(* Logix 5000 project; controller FV vendor 1 type 14 code 217 rev 31.11; software revision 31.00; part 12 of 63 *)
(* tags used below, declared in another part *)
   CWD : CHECKWORD_FLAGS;
   FR_B240 : INT[255];   // DEBOUNCE Debounce Flags
   FR_B246 : INT[255];   // V_REVERSE Flags for reversing contol action
   FR_B3 : INT[255];   // BINARY
   FR_FV26_AV07 : PlantItem;   // FV26_AV07
   FR_FV26_ROTO : PlantItem;   // FV26_ROTO
   FR_FV27_AV01 : PlantItem;   // FV27_AV01
   FR_FV27_AV04 : PlantItem;   // FV27_AV04
   FR_FV27_AV05 : PlantItem;   // FV27_AV05
   FR_FV27_AV06 : PlantItem;   // FV27_AV06
   FR_FV27_AV07 : PlantItem;   // FV27_AV07
   FR_FV27_ROTO : PlantItem;   // FV27_ROTO
   FR_FV27_VA01 : PlantItem;   // FV27_VA01
   FR_FV28_AV01 : PlantItem;   // FV28_AV01
   FR_FV28_AV04 : PlantItem;   // FV28_AV04
   FR_FV28_AV05 : PlantItem;   // FV28_AV05
   FR_FV28_AV06 : PlantItem;   // FV28_AV06
   FR_FV28_AV07 : PlantItem;   // FV28_AV07
   FR_FV28_ROTO : PlantItem;   // FV28_ROTO
   FR_FV28_V : PlantItem;   // FV28_V
   FR_FV28_VA01 : PlantItem;   // FV28_VA01
   FR_N10 : INT[265];   // FV_AGING Comms to FV Aging PL C
   FR_N100 : INT[265];   // FV FILLING
   FR_N110 : INT[265];   // GREEN BEER Green Beer Main
   FR_N120 : INT[265];   // YEAST CROP Yeast Cropping Main
   FR_N13 : INT[265];   // MV_ROUTE Comms to MV Routing PLC
   FR_N130 : INT[265];   // FILTRATE Filtrate Return
   FR_N14 : INT[265];   // MVFV CIP Comms to MVFV CIP Un it PLC
   FR_N160 : INT[265];   // VESSEL Vessel Working Direc tory
   FR_N200 : INT[265];   // ANALOG_IN Analog Inputs
   FR_N255 : INT[265];   // CHECKWORDS
   FR_N26 : INT[265];   // FV26
   FR_N27 : INT[265];   // FV27
   FR_N28 : INT[265];   // FV28
   FR_N7 : INT[265];   // INTEGER
   FR_N99 : INT[265];   // COMMENT Comment Lines
   FR_T144 : TIMER[255];   // CIP
   FR_T4 : TIMER[255];   // TIMER
   FR_T50 : TIMER[52];
   FR_T51 : TIMER[52];
   FR_T52 : TIMER[52];
   FR_T53 : TIMER[52];
   FR_VB1_AV08 : PlantItem;   // VB1_AV08
   FR_VB1_AV09 : PlantItem;   // VB1_AV09
   FR_VB2_AV04 : PlantItem;   // VB2_AV04
   FR_VB2_AV05 : PlantItem;   // VB2_AV05
   FR_VB4_AV02 : PlantItem;   // VB4_AV02
   FR_VB4_AV06 : PlantItem;   // VB4_AV06
   FR_VB4_AV08 : PlantItem;   // VB4_AV08
   FR_VB4_AV12 : PlantItem;   // VB4_AV12
   FR_VB4_AV14 : PlantItem;   // VB4_AV14
   FR_VB4_AV18 : PlantItem;   // VB4_AV18
(* FR_Common, continued *)

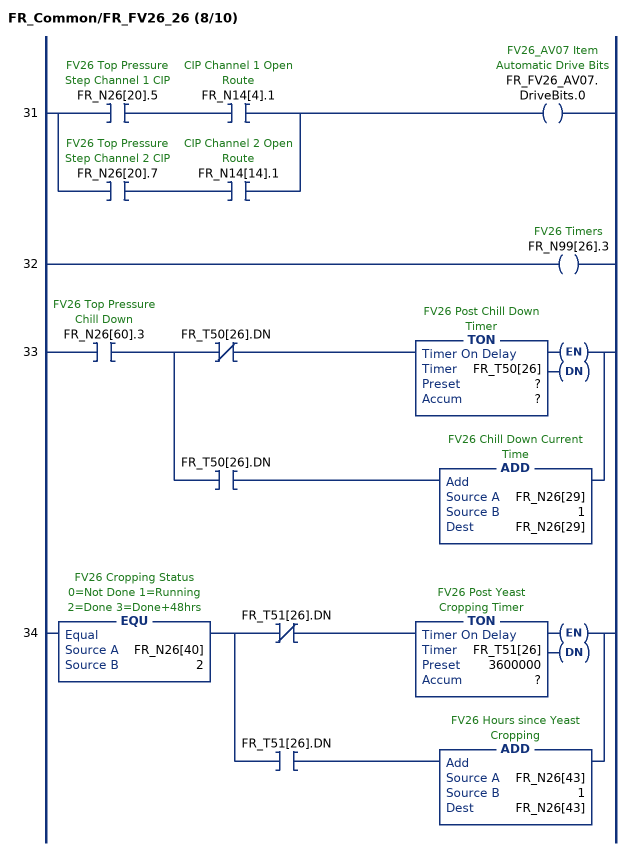
   [picture p160: FR_Common/FR_FV26_26 rungs 31-34]
   31: [XIC(FR_N26[20].5) XIC(FR_N14[4].1) ,XIC(FR_N26[20].7) XIC(FR_N14[14].1) ]OTE(FR_FV26_AV07.DriveBits.0);
   32: OTE(FR_N99[26].3);
   33: XIC(FR_N26[60].3)[XIO(FR_T50[26].DN) TON(FR_T50[26],?,?) ,XIC(FR_T50[26].DN) ADD(FR_N26[29],1,FR_N26[29]) ];
   34: EQU(FR_N26[40],2)[XIO(FR_T51[26].DN) TON(FR_T51[26],?,?) ,XIC(FR_T51[26].DN) ADD(FR_N26[43],1,FR_N26[43]) ];
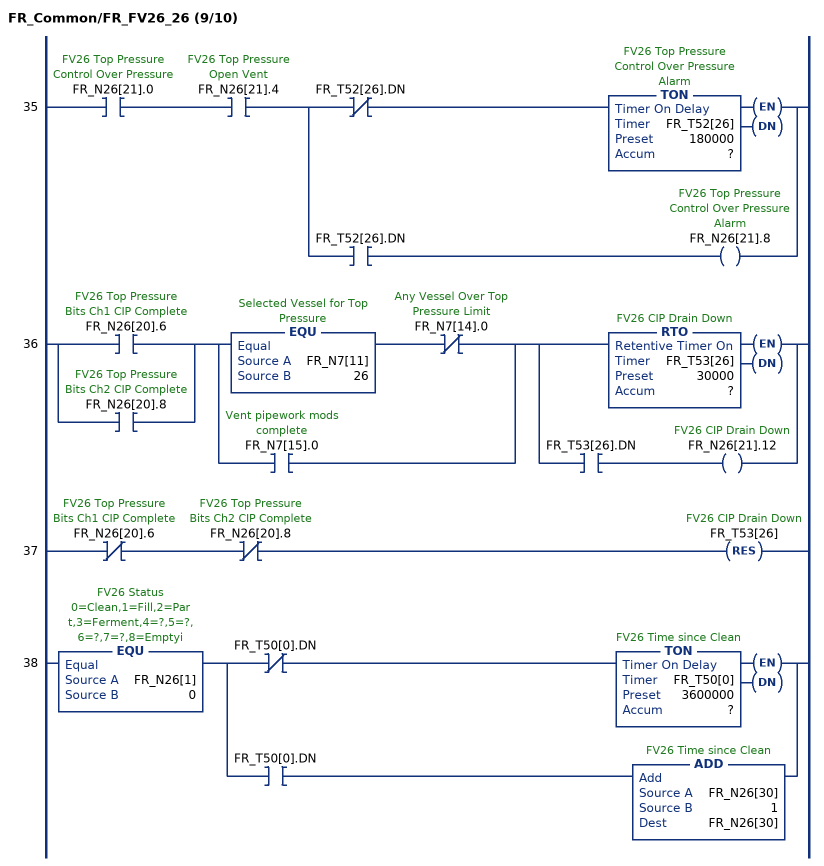
   35: XIC(FR_N26[21].0)XIC(FR_N26[21].4)[XIO(FR_T52[26].DN) TON(FR_T52[26],?,?) ,XIC(FR_T52[26].DN) OTE(FR_N26[21].8) ];
   36: [XIC(FR_N26[20].6) ,XIC(FR_N26[20].8) ][EQU(FR_N7[11],26) XIO(FR_N7[14].0) ,XIC(FR_N7[15].0) ][RTO(FR_T53[26],?,?) ,XIC(FR_T53[26].DN) OTE(FR_N26[21].12) ];
   37: XIO(FR_N26[20].6)XIO(FR_N26[20].8)RES(FR_T53[26]);
   38: EQU(FR_N26[1],0)[XIO(FR_T50[0].DN) TON(FR_T50[0],?,?) ,XIC(FR_T50[0].DN) ADD(FR_N26[30],1,FR_N26[30]) ];
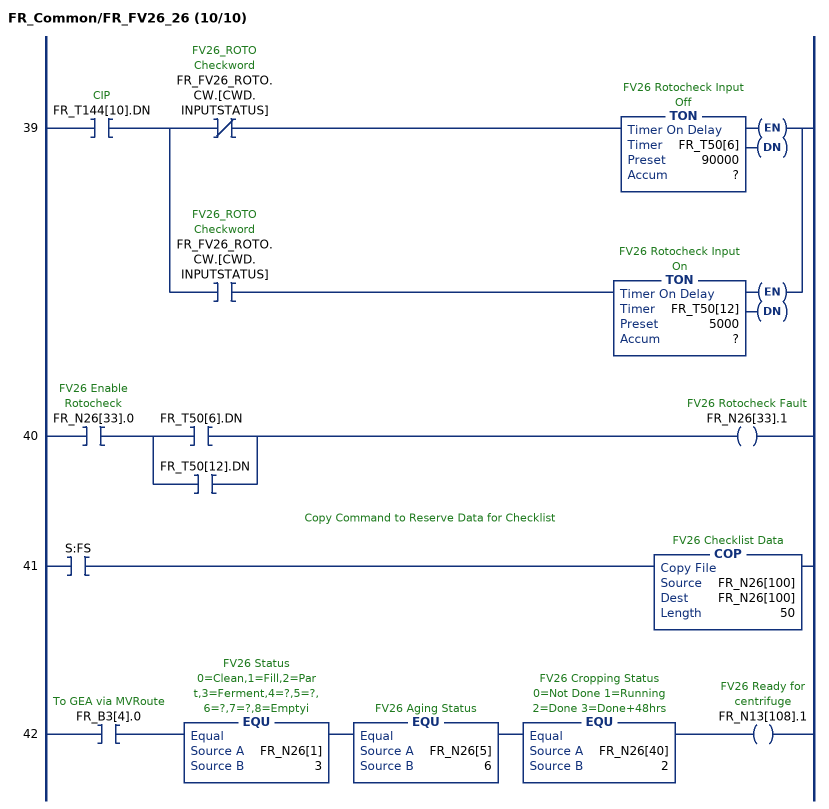
   39: XIC(FR_T144[10].DN)[XIO(FR_FV26_ROTO.CW.[CWD.INPUTSTATUS]) TON(FR_T50[6],?,?) ,XIC(FR_FV26_ROTO.CW.[CWD.INPUTSTATUS]) TON(FR_T50[12],?,?) ];
   40: XIC(FR_N26[33].0)[XIC(FR_T50[6].DN) ,XIC(FR_T50[12].DN) ]OTE(FR_N26[33].1);
   // Copy Command to Reserve Data for Checklist
   41: XIC(S:FS)COP(FR_N26[100],FR_N26[100],50);
   42: XIC(FR_B3[4].0)EQU(FR_N26[1],3)EQU(FR_N26[5],6)EQU(FR_N26[40],2)OTE(FR_N13[108].1);
END_ROUTINE

ROUTINE FR_FV27_27   (* ladder *)
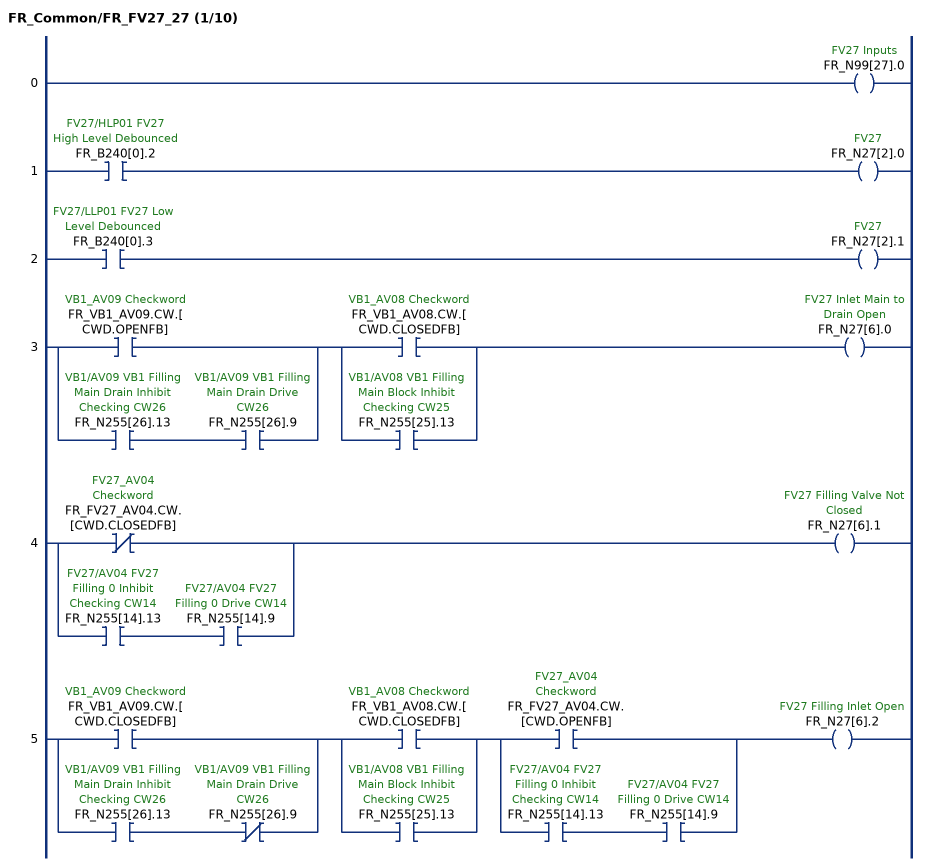
   0: OTE(FR_N99[27].0);
   1: XIC(FR_B240[0].2)OTE(FR_N27[2].0);
   2: XIC(FR_B240[0].3)OTE(FR_N27[2].1);
   3: [XIC(FR_VB1_AV09.CW.[CWD.OPENFB]) ,XIC(FR_N255[26].13) XIC(FR_N255[26].9) ][XIC(FR_VB1_AV08.CW.[CWD.CLOSEDFB]) ,XIC(FR_N255[25].13) ]OTE(FR_N27[6].0);
   4: [XIO(FR_FV27_AV04.CW.[CWD.CLOSEDFB]) ,XIC(FR_N255[14].13) XIC(FR_N255[14].9) ]OTE(FR_N27[6].1);
   5: [XIC(FR_VB1_AV09.CW.[CWD.CLOSEDFB]) ,XIC(FR_N255[26].13) XIO(FR_N255[26].9) ][XIC(FR_VB1_AV08.CW.[CWD.CLOSEDFB]) ,XIC(FR_N255[25].13) ][XIC(FR_FV27_AV04.CW.[CWD.OPENFB]) ,XIC(FR_N255[14].13) XIC(FR_N255[14].9) ]OTE(FR_N27[6].2);
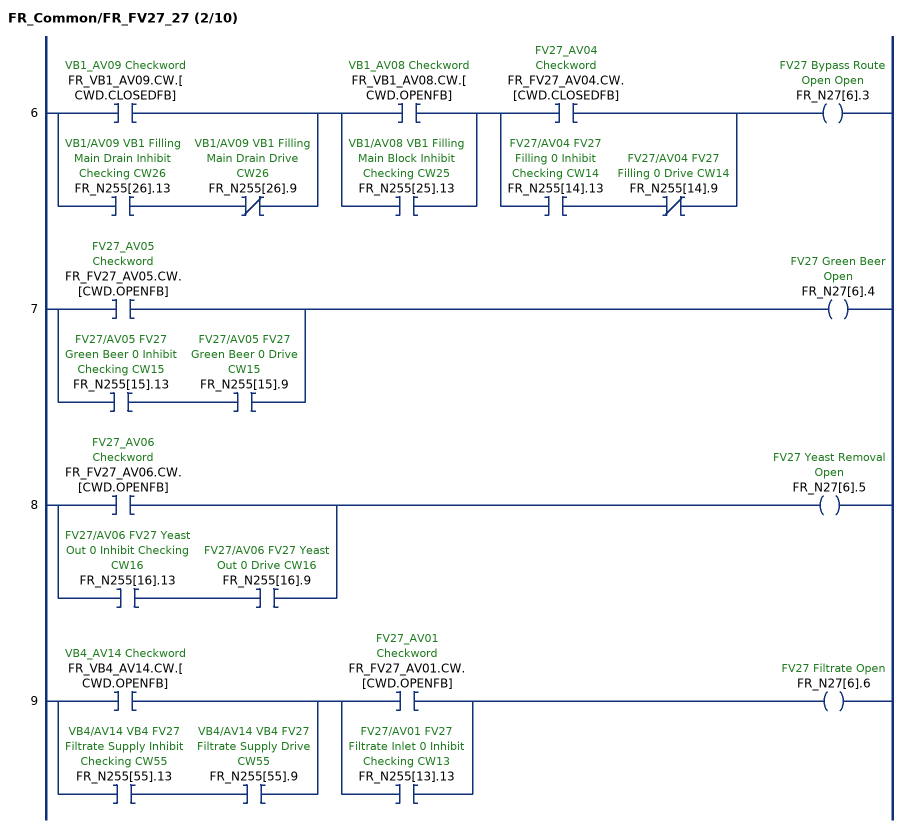
   6: [XIC(FR_VB1_AV09.CW.[CWD.CLOSEDFB]) ,XIC(FR_N255[26].13) XIO(FR_N255[26].9) ][XIC(FR_VB1_AV08.CW.[CWD.OPENFB]) ,XIC(FR_N255[25].13) ][XIC(FR_FV27_AV04.CW.[CWD.CLOSEDFB]) ,XIC(FR_N255[14].13) XIO(FR_N255[14].9) ]OTE(FR_N27[6].3);
   7: [XIC(FR_FV27_AV05.CW.[CWD.OPENFB]) ,XIC(FR_N255[15].13) XIC(FR_N255[15].9) ]OTE(FR_N27[6].4);
   8: [XIC(FR_FV27_AV06.CW.[CWD.OPENFB]) ,XIC(FR_N255[16].13) XIC(FR_N255[16].9) ]OTE(FR_N27[6].5);
   9: [XIC(FR_VB4_AV14.CW.[CWD.OPENFB]) ,XIC(FR_N255[55].13) XIC(FR_N255[55].9) ][XIC(FR_FV27_AV01.CW.[CWD.OPENFB]) ,XIC(FR_N255[13].13) ]OTE(FR_N27[6].6);
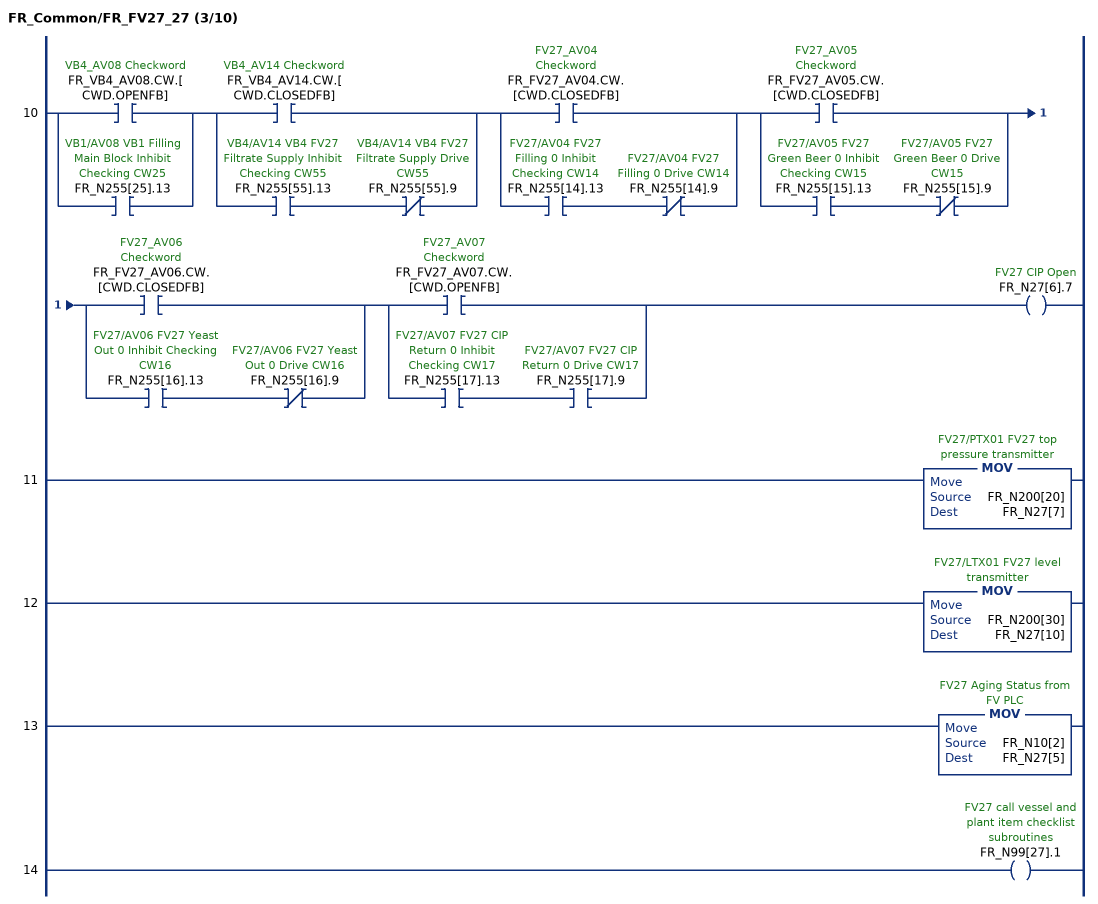
   10: [XIC(FR_VB4_AV08.CW.[CWD.OPENFB]) ,XIC(FR_N255[25].13) ][XIC(FR_VB4_AV14.CW.[CWD.CLOSEDFB]) ,XIC(FR_N255[55].13) XIO(FR_N255[55].9) ][XIC(FR_FV27_AV04.CW.[CWD.CLOSEDFB]) ,XIC(FR_N255[14].13) XIO(FR_N255[14].9) ][XIC(FR_FV27_AV05.CW.[CWD.CLOSEDFB]) ,XIC(FR_N255[15].13) XIO(FR_N255[15].9) ][XIC(FR_FV27_AV06.CW.[CWD.CLOSEDFB]) ,XIC(FR_N255[16].13) XIO(FR_N255[16].9) ][XIC(FR_FV27_AV07.CW.[CWD.OPENFB]) ,XIC(FR_N255[17].13) XIC(FR_N255[17].9) ]OTE(FR_N27[6].7);
   11: MOV(FR_N200[20],FR_N27[7]);
   12: MOV(FR_N200[30],FR_N27[10]);
   13: MOV(FR_N10[2],FR_N27[5]);
   14: OTE(FR_N99[27].1);
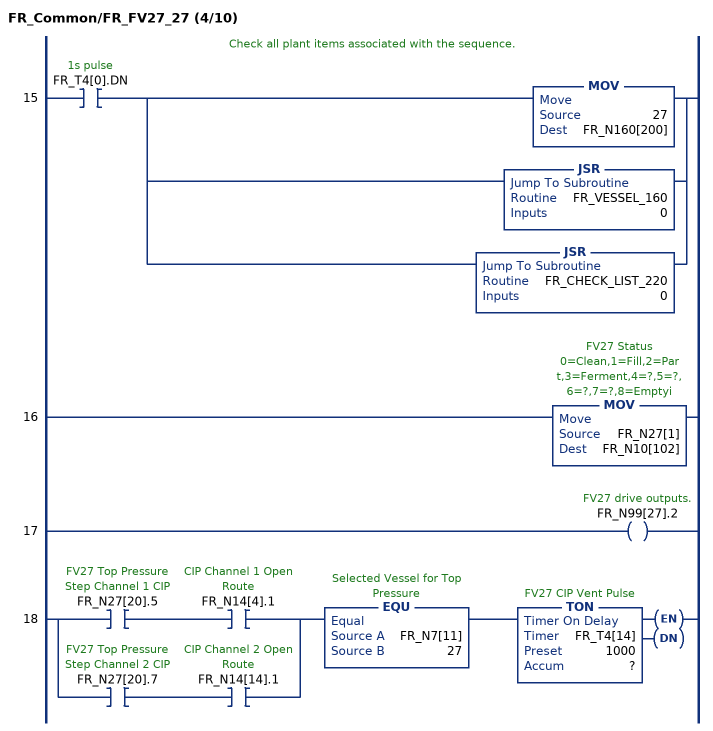
   // Check all plant items associated with the sequence.
   15: XIC(FR_T4[0].DN)[MOV(27,FR_N160[200]) ,JSR(FR_VESSEL_160,0) ,JSR(FR_CHECK_LIST_220,0) ];
   16: MOV(FR_N27[1],FR_N10[102]);
   17: OTE(FR_N99[27].2);
   18: [XIC(FR_N27[20].5) XIC(FR_N14[4].1) ,XIC(FR_N27[20].7) XIC(FR_N14[14].1) ]EQU(FR_N7[11],27)TON(FR_T4[14],?,?);
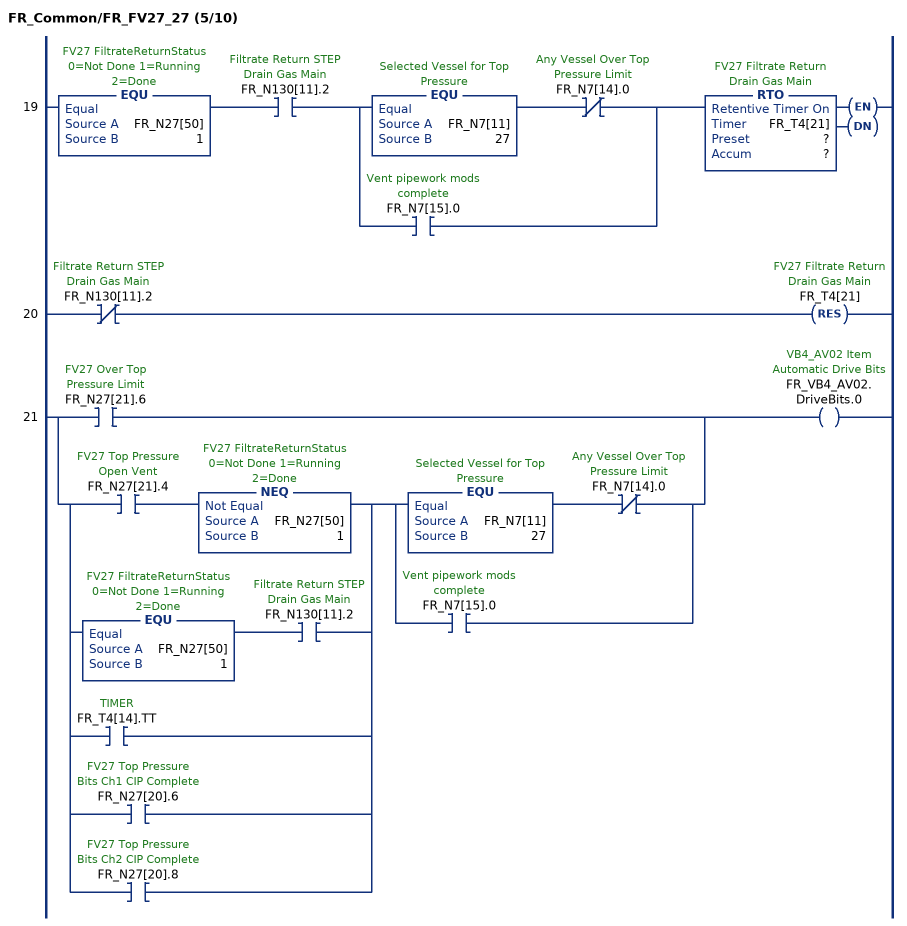
   19: EQU(FR_N27[50],1)XIC(FR_N130[11].2)[EQU(FR_N7[11],27) XIO(FR_N7[14].0) ,XIC(FR_N7[15].0) ]RTO(FR_T4[21],?,?);
   20: XIO(FR_N130[11].2)RES(FR_T4[21]);
   21: [XIC(FR_N27[21].6) ,[XIC(FR_N27[21].4) NEQ(FR_N27[50],1) ,EQU(FR_N27[50],1) XIC(FR_N130[11].2) ,XIC(FR_T4[14].TT) ,[XIC(FR_N27[20].6) ,XIC(FR_N27[20].8) ] ] [EQU(FR_N7[11],27) XIO(FR_N7[14].0) ,XIC(FR_N7[15].0) ] ]OTE(FR_VB4_AV02.DriveBits.0);
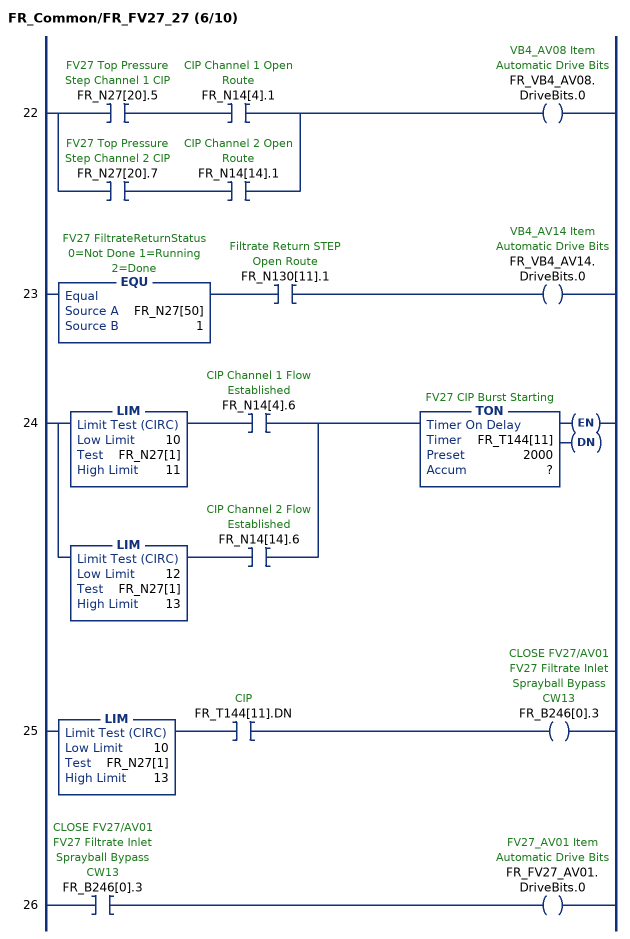
   22: [XIC(FR_N27[20].5) XIC(FR_N14[4].1) ,XIC(FR_N27[20].7) XIC(FR_N14[14].1) ]OTE(FR_VB4_AV08.DriveBits.0);
   23: EQU(FR_N27[50],1)XIC(FR_N130[11].1)OTE(FR_VB4_AV14.DriveBits.0);
   24: [LIM(10,FR_N27[1],11) XIC(FR_N14[4].6) ,LIM(12,FR_N27[1],13) XIC(FR_N14[14].6) ]TON(FR_T144[11],?,?);
   25: LIM(10,FR_N27[1],13)XIC(FR_T144[11].DN)OTE(FR_B246[0].3);
   26: XIC(FR_B246[0].3)OTE(FR_FV27_AV01.DriveBits.0);
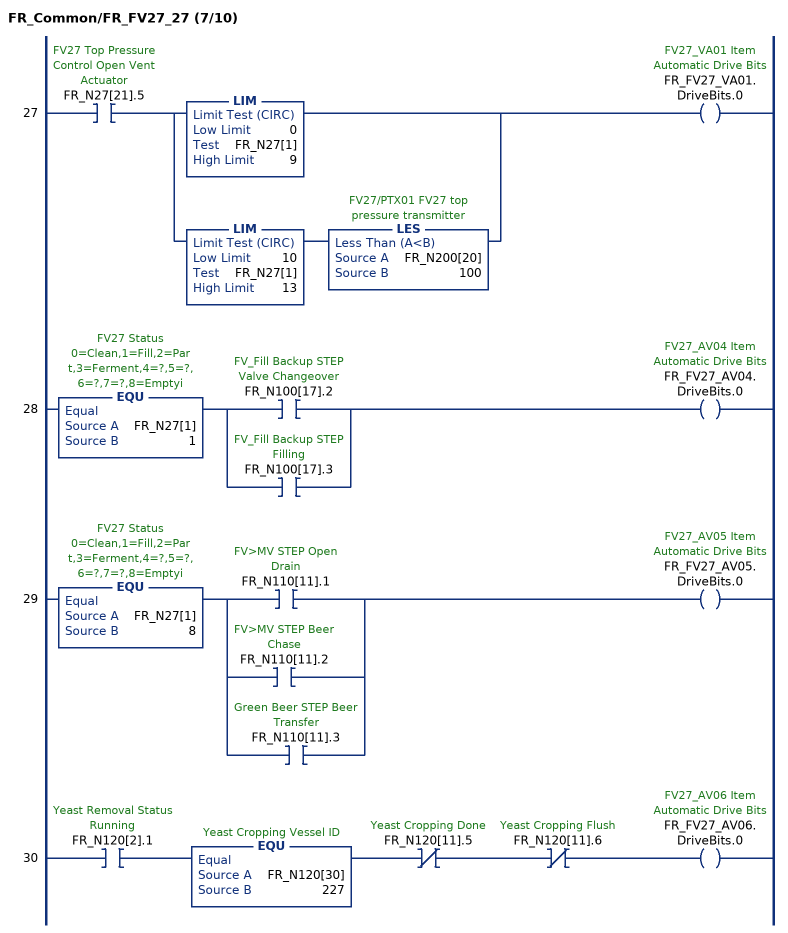
   27: XIC(FR_N27[21].5)[LIM(0,FR_N27[1],9) ,LIM(10,FR_N27[1],13) LES(FR_N200[20],100) ]OTE(FR_FV27_VA01.DriveBits.0);
   28: EQU(FR_N27[1],1)[XIC(FR_N100[17].2) ,XIC(FR_N100[17].3) ]OTE(FR_FV27_AV04.DriveBits.0);
   29: EQU(FR_N27[1],8)[XIC(FR_N110[11].1) ,XIC(FR_N110[11].2) ,XIC(FR_N110[11].3) ]OTE(FR_FV27_AV05.DriveBits.0);
   30: XIC(FR_N120[2].1)EQU(FR_N120[30],227)XIO(FR_N120[11].5)XIO(FR_N120[11].6)OTE(FR_FV27_AV06.DriveBits.0);
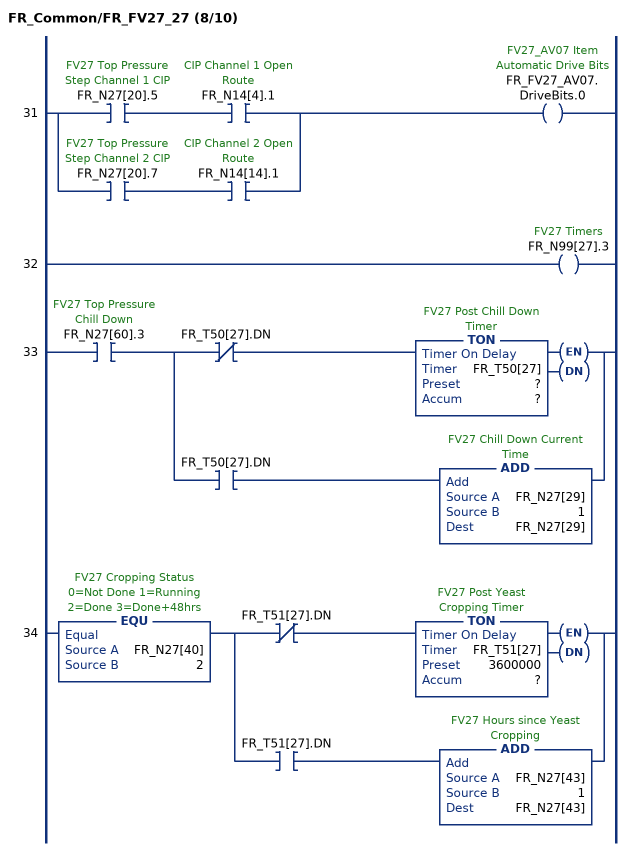
   31: [XIC(FR_N27[20].5) XIC(FR_N14[4].1) ,XIC(FR_N27[20].7) XIC(FR_N14[14].1) ]OTE(FR_FV27_AV07.DriveBits.0);
   32: OTE(FR_N99[27].3);
   33: XIC(FR_N27[60].3)[XIO(FR_T50[27].DN) TON(FR_T50[27],?,?) ,XIC(FR_T50[27].DN) ADD(FR_N27[29],1,FR_N27[29]) ];
   34: EQU(FR_N27[40],2)[XIO(FR_T51[27].DN) TON(FR_T51[27],?,?) ,XIC(FR_T51[27].DN) ADD(FR_N27[43],1,FR_N27[43]) ];